
screen "BWTS" 480x228, template "Template_1"
   on GenerateScreen: "TitleUpdater"()
   GraphicView "Graphic view_6" at 70,107 size 332x4; Picture "Graphic_151"
   Button "Button_2" at 88,1 size 50x40; TextOff 'IGGS'
      on Release: ActivateScreen("IGGS Plant", 0)
   Button "Button_4" at 144,1 size 50x40; TextOff 'PGC'
      on Release: ActivateScreen("PGC", 0)
   Button "Button_6" at 199,2 size 50x40; TextOff 'GCU'
      on Release: ActivateScreen("GCU Plant", 0)
   Button "Button_1" at 88,1 size 50x40; TextOff 'IGGS'
      on Release: ActivateScreen("IGGS Plant", 0)
      Visibility <- "IGG Running"
   Button "Button_3" at 144,1 size 50x40; TextOff 'PGC'
      on Release: ActivateScreen("PGC", 0)
      Visibility <- "Process Gas Compressor Running/Stopped"
   Button "Button_5" at 199,2 size 50x40; TextOff 'GCU'
      on Release: ActivateScreen("GCU Plant", 0)
      Visibility <- "100_GCU_AUTO_SEQ_DB_CRNT_STEP"
   Button "HmiScreenItemData_2" at 364,2 size 115x30; TextOn 'I&A Compressor Ok'; TextOff 'Previous Screen'
      on Release: function_efd93a16()
   Button "HmiScreenItemData_19" at 270,2 size 85x40; TextOn 'IGG Plant'; TextOff 'Alarms'
      on Release: ActivateScreen("Alarms", 0)
   Button "Button_20" at 205,191 size 60x34; TextOff 'Dwell'
      Appearance <- "2100_BTCS_CNTRL_DB_BTCS_STATE"
   Button "Button_21" at 2,191 size 60x34; TextOff 'Un- selected'
      Appearance <- "HMI Indication Logic_DB_Tank Selected"
   Button "Button_22" at 69,191 size 60x34; TextOff 'Selected'
      Appearance <- "HMI Indication Logic_DB_Tank Selected"
   Button "Button_23" at 137,191 size 60x34; TextOff 'De-Oxy'
      Appearance <- "2100_BTCS_CNTRL_DB_BTCS_STEP"
   Button "Button_24" at 272,191 size 60x34; TextOff 'Re-Oxy'
      Appearance <- "2100_BTCS_CNTRL_DB_BTCS_STEP"
   Button "Button_25" at 340,191 size 60x34; TextOff 'Post Dwell'
      Appearance <- "2100_BTCS_CNTRL_DB_BTCS_STATE"
   Button "Button_26" at 408,191 size 70x34; TextOff 'Complete'
      Appearance <- "HMI Indication Logic_DB_Sequence Finished"
   TextField "Text field_1" at 185,171 size 116x21; Text 'TANK STATUS'
   Button "Button_28" at 80,49 size 50x55; TextOff 'Tank 6P'
      on Release: function_efd93a16("Tank 6S Status", 0, 0, -1, 2, 1)
   Button "Button_13" at 80,49 size 50x55; TextOff 'Tank 6P'
      on Release: function_efd93a16("Tank 6S Status", 0, 0, -1, 2, 1)
      Appearance <- "2100_BTCS_CNTRL_DB_BTCS_STATE"
      Visibility <- "504_Tank Grouping_DB2020_GROUP of TANK 12"
   Button "Button_29" at 132,49 size 50x55; TextOff 'Tank 5P'
      on Release: function_efd93a16("Tank 5S Status", 0, 0, -1, 2, 1)
   Button "Button_12" at 132,49 size 50x55; TextOff 'Tank 5P'
      on Release: function_efd93a16("Tank 5S Status", 0, 0, -1, 2, 1)
      Appearance <- "2100_BTCS_CNTRL_DB_BTCS_STATE"
      Visibility <- "504_Tank Grouping_DB2020_GROUP of TANK 10"
   Button "Button_30" at 185,49 size 50x55; TextOff 'Tank 4P'
      on Release: function_efd93a16("Tank 4S Status", 0, 0, -1, 2, 1)
   Button "Button_15" at 185,49 size 50x55; TextOff 'Tank 4P'
      on Release: function_efd93a16("Tank 4S Status", 0, 0, -1, 2, 1)
      Appearance <- "2100_BTCS_CNTRL_DB_BTCS_STATE"
      Visibility <- "504_Tank Grouping_DB2020_GROUP of TANK 8"
   Button "Button_31" at 238,49 size 50x55; TextOff 'Tank 3P'
      on Release: function_efd93a16("Tank 3S Status", 0, 0, -1, 2, 1)
   Button "Button_14" at 238,49 size 50x55; TextOff 'Tank 3P'
      on Release: function_efd93a16("Tank 3S Status", 0, 0, -1, 2, 1)
      Appearance <- "2100_BTCS_CNTRL_DB_BTCS_STATE"
      Visibility <- "504_Tank Grouping_DB2020_GROUP of TANK 6"
   Button "Button_32" at 291,49 size 50x55; TextOff 'Tank 2P'
      on Release: function_efd93a16("Tank 2S Status", 0, 0, -1, 2, 1)
   Button "Button_17" at 291,49 size 50x55; TextOff 'Tank 2P'
      on Release: function_efd93a16("Tank 2S Status", 0, 0, -1, 2, 1)
      Appearance <- "2100_BTCS_CNTRL_DB_BTCS_STATE"
      Visibility <- "504_Tank Grouping_DB2020_GROUP of TANK 4"
   Button "Button_33" at 344,49 size 50x55; TextOff 'Tank 1P'
      on Release: function_efd93a16("Tank 1S Status", 0, 0, -1, 2, 1)
   Button "Button_16" at 344,49 size 50x55; TextOff 'Tank 1P'
      on Release: function_efd93a16("Tank 1S Status", 0, 0, -1, 2, 1)
      Appearance <- "2100_BTCS_CNTRL_DB_BTCS_STATE"
      Visibility <- "504_Tank Grouping_DB2020_GROUP of TANK 2"
   Button "Button_34" at 402,82 size 50x55; TextOff 'FP Tank'
      on Release: function_efd93a16("Tank FP Status", 0, 0, -1, 2, 1)
   Button "Button_19" at 402,82 size 50x55; TextOff 'FP Tank'
      on Release: function_efd93a16("Tank FP Status", 0, 0, -1, 2, 1)
      Appearance <- "2100_BTCS_CNTRL_DB_BTCS_STATE"
      Visibility <- "504_Tank Grouping_DB2020_GROUP of TANK 1"
   Button "Button_35" at 22,82 size 50x55; TextOff 'AP Tank'
      on Release: function_efd93a16("Tank AP Status", 0, 0, -1, 2, 1)
   Button "Button_18" at 22,82 size 50x55; TextOff 'AP Tank'
      on Release: function_efd93a16("Tank AP Status", 0, 0, -1, 2, 1)
      Appearance <- "2100_BTCS_CNTRL_DB_BTCS_STATE"
      Visibility <- "504_Tank Grouping_DB2020_GROUP of TANK 14"
   Button "Button_36" at 80,114 size 50x55; TextOff 'Tank 6S'
      on Release: function_efd93a16("Tank 6P Status", 0, 0, -1, 2, 1)
   Button "Button_7" at 80,114 size 50x55; TextOff 'Tank 6S'
      on Release: function_efd93a16("Tank 6P Status", 0, 0, -1, 2, 1)
      Appearance <- "2100_BTCS_CNTRL_DB_BTCS_STATE"
      Visibility <- "504_Tank Grouping_DB2020_GROUP of TANK 13"
   Button "Button_37" at 132,114 size 50x55; TextOff 'Tank 5S'
      on Release: function_efd93a16("Tank 5P Status", 0, 0, -1, 2, 1)
   Button "Button_27" at 132,114 size 50x55; TextOff 'Tank 5S'
      on Release: function_efd93a16("Tank 5P Status", 0, 0, -1, 2, 1)
      Appearance <- "2100_BTCS_CNTRL_DB_BTCS_STATE"
      Visibility <- "504_Tank Grouping_DB2020_GROUP of TANK 11"
   Button "Button_38" at 185,114 size 50x55; TextOff 'Tank 4S'
      on Release: function_efd93a16("Tank 4P Status", 0, 0, -1, 2, 1)
   Button "Button_9" at 185,114 size 50x55; TextOff 'Tank 4S'
      on Release: function_efd93a16("Tank 4P Status", 0, 0, -1, 2, 1)
      Appearance <- "2100_BTCS_CNTRL_DB_BTCS_STATE"
      Visibility <- "504_Tank Grouping_DB2020_GROUP of TANK 9"
   Button "Button_39" at 238,114 size 50x55; TextOff 'Tank 3S'
      on Release: function_efd93a16("Tank 3P Status", 0, 0, -1, 2, 1)
   Button "Button_8" at 238,114 size 50x55; TextOff 'Tank 3S'
      on Release: function_efd93a16("Tank 3P Status", 0, 0, -1, 2, 1)
      Appearance <- "2100_BTCS_CNTRL_DB_BTCS_STATE"
      Visibility <- "504_Tank Grouping_DB2020_GROUP of TANK 7"
   Button "Button_40" at 291,114 size 50x55; TextOff 'Tank 2S'
      on Release: function_efd93a16("Tank 2P Status", 0, 0, -1, 2, 1)
   Button "Button_11" at 291,114 size 50x55; TextOff 'Tank 2S'
      on Release: function_efd93a16("Tank 2P Status", 0, 0, -1, 2, 1)
      Appearance <- "2100_BTCS_CNTRL_DB_BTCS_STATE"
      Visibility <- "504_Tank Grouping_DB2020_GROUP of TANK 5"
   Button "Button_41" at 344,114 size 50x55; TextOff 'Tank 1S'
      on Release: function_efd93a16("Tank 1P Status", 0, 0, -1, 2, 1)
   Button "Button_10" at 344,114 size 50x55; TextOff 'Tank 1S'
      on Release: function_efd93a16("Tank 1P Status", 0, 0, -1, 2, 1)
      Appearance <- "2100_BTCS_CNTRL_DB_BTCS_STATE"
      Visibility <- "504_Tank Grouping_DB2020_GROUP of TANK 3"
   Polyline "Polyline_1" at 80,49 size 48x54
      Visibility <- "504_Tank Grouping_DB2020_RUN TANK 12"
   Polyline "Polyline_2" at 80,114 size 48x54
      Visibility <- "504_Tank Grouping_DB2020_RUN TANK 13"
   Polyline "Polyline_3" at 133,114 size 48x54
      Visibility <- "504_Tank Grouping_DB2020_RUN TANK 11"
   Polyline "Polyline_4" at 132,49 size 48x54
      Visibility <- "504_Tank Grouping_DB2020_RUN TANK 10"
   Polyline "Polyline_5" at 185,49 size 48x54
      Visibility <- "504_Tank Grouping_DB2020_RUN TANK 8"
   Polyline "Polyline_6" at 185,114 size 48x54
      Visibility <- "504_Tank Grouping_DB2020_RUN TANK 9"
   Polyline "Polyline_7" at 239,49 size 48x54
      Visibility <- "504_Tank Grouping_DB2020_RUN TANK 6"
   Polyline "Polyline_8" at 238,114 size 48x54
      Visibility <- "504_Tank Grouping_DB2020_RUN TANK 7"
   Polyline "Polyline_9" at 292,114 size 48x54
      Visibility <- "504_Tank Grouping_DB2020_RUN TANK 5"
   Polyline "Polyline_10" at 291,49 size 48x54
      Visibility <- "504_Tank Grouping_DB2020_RUN TANK 4"
   Polyline "Polyline_11" at 345,49 size 48x54
      Visibility <- "504_Tank Grouping_DB2020_RUN TANK 2"
   Polyline "Polyline_12" at 345,114 size 48x54
      Visibility <- "504_Tank Grouping_DB2020_RUN TANK 3"
   Polyline "Polyline_13" at 403,82 size 48x54
      Visibility <- "504_Tank Grouping_DB2020_RUN TANK 1"
   Polyline "Polyline_14" at 22,82 size 48x54
      Visibility <- "504_Tank Grouping_DB2020_RUN TANK 14"
   Button "HmiScreenItemData_1" at 1,1 size 84x30; TextOn 'I&A Compressor Ok'; TextOff 'Main Index'
      on Release: ActivateScreen("Main Index", 0)

screen "PGC" 480x228, template "Template_1"
   on GenerateScreen: "TitleUpdater"()
   Button "HmiScreenItemData_6" at 353,1 size 126x30; TextOn 'I&A Compressor Ok'; TextOff 'Previous Screen'
      on Release: function_efd93a16()
   TextField "Text field_7" at 4,38 size 278x22; Text 'Process Gas Compressor Control'
   Button "Button_15" at 23,138 size 57x23; TextOn 'Enabled'; TextOff 'Disabled'
   Button "Button_16" at 177,138 size 64x23; TextOn 'Alarm'; TextOff 'Text'
   TextField "Text field_15" at 27,118 size 56x17; Text 'Enabled'
   TextField "Text field_16" at 102,118 size 58x17; Text 'Running'
   TextField "Text field_18" at 179,117 size 69x17; Text 'Shutdown'
   Button "Button_1" at 100,138 size 57x23; TextOn 'Enabled'; TextOff 'Stopped'
   TextField "Text field_32" at 23,139 size 57x23; Text 'Enabled'
      Visibility <- "10_DI_DATA_E_400_SHTDN"
   TextField "Text field_2" at 100,138 size 57x23; Text 'Running'
      Visibility <- "10_DI_DATA_E_400_RUN"
   Button "Button_2" at 177,138 size 64x23; TextOn 'Alarm'; TextOff 'Shutdown'
      Appearance <- "10_DI_DATA_E_400_NOK"
      Visibility <- "10_DI_DATA_E_400_NOK"
   Button "Button_7" at 262,38 size 57x23; TextOn 'Alarm'; TextOff 'Service'
      Appearance <- "140_PGC_HRS_RUN_DB_SRVC"
   GraphicView "Graphic view_1" at 288,29 size 192x199; Picture "Graphic_251"
   Button "HmiScreenItemData_1" at 1,1 size 84x30; TextOn 'I&A Compressor Ok'; TextOff 'Main Index'
      on Release: ActivateScreen("Main Index", 0)

screen "CA Blower" 480x228, template "Template_1"
   on GenerateScreen: "TitleUpdater"()
   Button "HmiScreenItemData_6" at 353,1 size 126x30; TextOn 'I&A Compressor Ok'; TextOff 'Previous Screen'
      on Release: function_efd93a16()
   GraphicIOField "Graphic I/O field_2" at 281,42 size 196x184; PictureList "IA Compressor"
      ProcessValue <- "CA Blower Animation"
   Button "Button_3" at 126,118 size 57x23; TextOn 'Enabled'; TextOff 'Disabled'
   TextField "Text field_4" at 129,98 size 56x17; Text 'Enabled'
   TextField "Text field_5" at 202,98 size 38x17; Text 'Fault'
   Button "Button_5" at 192,118 size 57x23; TextOn 'Enabled'; TextOff 'Healthy'
   TextField "Text field_8" at 126,118 size 57x23; Text 'Enabled'
      Visibility <- "CA Blower Control"
   Button "Button_6" at 192,118 size 57x23; TextOn 'Alarm'; TextOff 'Fault'
      Visibility <- "Data To IGG PLC_Data_VSD Fault Flag"
      Appearance <- "Data To IGG PLC_Data_VSD Fault Flag"
   TextField "Text field_3" at 5,120 size 119x18; Text 'Combustion Air'
   TextField "Text field_7" at 4,38 size 263x22; Text 'Combustion Air Blower Control'
   Button "Button_7" at 276,38 size 57x23; TextOn 'Alarm'; TextOff 'Service'
      Appearance <- "Operation hours E139_IDB_Service Time bit"
   Button "HmiScreenItemData_1" at 1,1 size 84x30; TextOn 'I&A Compressor Ok'; TextOff 'Main Index'
      on Release: ActivateScreen("Main Index", 0)

screen "Cooling System" 480x228, template "Template_1"
   on GenerateScreen: "TitleUpdater"()
   Button "HmiScreenItemData_6" at 353,1 size 126x30; TextOn 'I&A Compressor Ok'; TextOff 'Previous Screen'
      on Release: function_efd93a16()
   TextField "Text field_7" at 140,69 size 201x22; Text 'Cooling System Control'
   Button "Button_15" at 207,128 size 57x23; TextOn 'Enabled'; TextOff 'Disabled'
   Button "Button_16" at 361,128 size 64x23; TextOn 'Alarm'; TextOff 'Text'
   TextField "Text field_14" at 35,130 size 179x18; Text 'Cooling Sea Water Pump'
   TextField "Text field_15" at 211,108 size 56x17; Text 'Enabled'
   TextField "Text field_16" at 286,108 size 58x17; Text 'Running'
   TextField "Text field_18" at 363,107 size 69x17; Text 'Shutdown'
   Rectangle "Rectangle_10" at 33,123 size 166x32
      Appearance <- "P301 Present"
   Button "Button_1" at 284,128 size 57x23; TextOn 'Enabled'; TextOff 'Stopped'
   TextField "Text field_32" at 207,128 size 57x23; Text 'Enabled'
      Visibility <- "CSW Pump Enabled"
   TextField "Text field_2" at 284,128 size 57x23; Text 'Running'
      Visibility <- "Data_To_BC PLC_Data_Cooling Water System Proved"
   Button "Button_2" at 361,128 size 64x23; TextOn 'Alarm'; TextOff 'Shutdown'
      Visibility <- "Cooling Sea Water Pump Shutdown"
      Appearance <- "Cooling Sea Water Pump Shutdown"
   Rectangle "Rectangle_1" at 24,99 size 425x69
      Visibility <- "P301 Present"
   Group "Group" at 15,161 size 490x34
   Button "HmiScreenItemData_1" at 1,1 size 84x30; TextOn 'I&A Compressor Ok'; TextOff 'Main Index'
      on Release: ActivateScreen("Main Index", 0)
   TextField "Text field_1" at 28,161 size 466x34; Text 'Cooling System Pressure in Range'
      Visibility <- "Cooling System Operating"
   TextField "Text field_3" at 15,162 size 490x32; Text 'Cooling System Pressure Out of Range'
      Visibility <- "Cooling System Operating"

screen "Fuel System" 480x228, template "Template_1"
   on GenerateScreen: "TitleUpdater"()
   Button "HmiScreenItemData_6" at 172,1 size 126x30; TextOn 'I&A Compressor Ok'; TextOff 'Previous Screen'
      on Release: function_efd93a16()
   GraphicView "Graphic view_4" at 271,104 size 24x23; Picture "Graphic_102"
   TextField "Text field_3" at 359,196 size 55x18; Text 'E-500B'
   GraphicView "Graphic view_16" at 326,49 size 123x15; Picture "Graphic_99"
   GraphicIOField "Graphic I/O field_1" at 354,30 size 60x65; PictureList "Pump Ani"
      ProcessValue <- "Fuel Pump 1 Animation"
   GraphicView "Graphic view_10" at 325,151 size 124x15; Picture "Graphic_99"
   GraphicIOField "Graphic I/O field_2" at 354,133 size 60x65; PictureList "Pump Ani"
      ProcessValue <- "Fuel Pump 2 Animation"
   GraphicView "Graphic view_17" at 310,64 size 15x94; Picture "Graphic_101"
   GraphicView "Graphic view_14" at 311,140 size 21x25; Picture "Graphic_96"
   GraphicView "Graphic view_18" at 311,50 size 24x23; Picture "Graphic_102"
   GraphicView "Graphic view_19" at 306,99 size 18x23; Picture "Graphic_105"
   GraphicView "Graphic view_20" at 450,64 size 15x94; Picture "Graphic_101"
   GraphicView "Graphic view_9" at 440,50 size 24x23; Picture "Graphic_104"
   GraphicView "Graphic view_21" at 439,141 size 25x24; Picture "Graphic_97"
   GraphicView "Graphic view_7" at 451,100 size 19x24; Picture "Graphic_103"
   GraphicView "Graphic view_22" at 296,103 size 9x15; Picture "Graphic_99"
   GraphicView "Graphic view_24" at 340,49 size 18x15; Picture "Graphic_99"
   TextField "Text field_2" at 359,96 size 56x18; Text 'E-500A'
   GraphicView "Graphic view_1" at 289,103 size 27x15; Picture "Graphic_99"
   Rectangle "Rectangle_13" at 346,24 size 77x92
      Appearance <- "Fuel Pump 1 Tripped"
   Rectangle "Rectangle_14" at 346,127 size 77x92
      Appearance <- "Fuel Pump 2 Tripped"
   TextField "Text field_7" at 334,225 size 83x18; Text 'Duty Pump'
      Visibility <- "101_Fuel_Pumps_DB_Duty Is B"
   TextField "Text field_12" at 346,7 size 83x18; Text 'Duty Pump'
      Visibility <- "101_Fuel_Pumps_DB_Duty Is A"
   Button "HmiScreenItemData_7" at 209,128 size 84x37; TextOn 'Back'; TextOff 'PSelect'; Authorization "Operate"
      on Press: function_b14e0dd5("HMI Fuel Pump Duty Select", 0)
   Button "Button_15" at 7,61 size 57x25; TextOn 'Enabled'; TextOff 'Disabled'
   TextField "Text field_14" at 1,92 size 92x20; Text 'Fuel Pump 1'
   TextField "Text field_15" at 11,40 size 60x18; Text 'Enabled'
   Button "Button_17" at 229,61 size 57x25; TextOn 'Alarm'; TextOff 'Service'
   Button "Button_9" at 229,61 size 57x25; TextOn 'Alarm'; TextOff 'Service'
      Visibility <- "82_To_HMI_E500A Fuel Pump Service Due"
   Button "Button_13" at 7,61 size 57x25; TextOn 'Enabled'; TextOff 'Enabled'
      Visibility <- "Fuel Pump 1 Enabled"
   IOField "I/O field_3" at 131,61 size 65x25; FormatPattern 999999
      ProcessValue <- "64_Functioning Hours_E500A_IDB_Hours Functioning"
   TextField "Text field_5" at 131,38 size 72x18; Text 'Hour Run'
   Button "Button_1" at 70,61 size 57x25; TextOn 'Alarm'; TextOff 'Text'
   TextField "Text field_6" at 78,38 size 45x18; Text 'Alarm'
   Button "Button_3" at 70,61 size 57x25; TextOn 'Alarm'; TextOff 'Tripped'
      Visibility <- "Fuel Pump 1 Tripped"
      Appearance <- "Fuel Pump 1 Tripped"
   Button "Button_18" at 7,178 size 57x25; TextOn 'Enabled'; TextOff 'Disabled'
   TextField "Text field_19" at 1,208 size 92x20; Text 'Fuel Pump 2'
   Button "Button_20" at 229,178 size 57x25; TextOn 'Alarm'; TextOff 'Service'
   Button "Button_10" at 229,178 size 57x25; TextOn 'Alarm'; TextOff 'Service'
      Visibility <- "82_To_HMI_E500B Fuel Pump Service Due"
   Button "Button_14" at 7,177 size 57x25; TextOn 'Enabled'; TextOff 'Enabled'
      Visibility <- "Fuel Pump 2 Enabled"
   IOField "I/O field_6" at 131,177 size 65x25; FormatPattern 999999
      ProcessValue <- "64_Functioning Hours_E500B_IDB_Hours Functioning"
   Button "Button_2" at 70,177 size 57x25; TextOn 'Alarm'; TextOff 'Text'
   Button "Button_4" at 70,177 size 57x25; TextOn 'Alarm'; TextOff 'Tripped'
      Visibility <- "Fuel Pump 2 Tripped"
      Appearance <- "Fuel Pump 2 Tripped"
   Button "HmiScreenItemData_1" at 1,1 size 84x30; TextOn 'I&A Compressor Ok'; TextOff 'Main Index'
      on Release: ActivateScreen("Main Index", 0)

screen "Alarms" 480x228, template "Template_1"
   on GenerateScreen: "TitleUpdater"()
   AlarmView "Alarm view_1" at 0,31 size 480x196
   Button "HmiScreenItemData_6" at 353,1 size 126x30; TextOn 'I&A Compressor Ok'; TextOff 'Previous Screen'
      on Release: function_efd93a16()
   Button "HmiScreenItemData_1" at 1,1 size 84x30; TextOn 'I&A Compressor Ok'; TextOff 'Main Index'
      on Release: ActivateScreen("Main Index", 0)

screen "Events History" 480x228, template "Template_1"
   on GenerateScreen: "TitleUpdater"()
   AlarmView "Alarm view_1" at 0,44 size 480x184
   Button "HmiScreenItemData_1" at 1,1 size 84x30; TextOn 'I&A Compressor Ok'; TextOff 'Main Index'
      on Release: ActivateScreen("Main Index", 0)

screen "Air System" 480x228, template "Template_1"
   on GenerateScreen: "TitleUpdater"()
   Button "HmiScreenItemData_6" at 353,1 size 126x30; TextOn 'I&A Compressor Ok'; TextOff 'Previous Screen'
      on Release: function_efd93a16()
   TextField "Text field_1" at 0,38 size 368x23; Text 'Instrument & Atomising Air Compressor'
   Button "Button_4" at 362,39 size 57x23; TextOn 'Alarm'; TextOff 'Service'
      Visibility <- "IDB_E131_Functioning Hours_Service Time bit"
      Appearance <- "IDB_E131_Functioning Hours_Service Time bit"
   Button "Button_15" at 27,137 size 57x23; TextOn 'Enabled'; TextOff 'Disabled'
   Button "Button_16" at 181,137 size 64x23; TextOn 'Alarm'; TextOff 'Text'
   TextField "Text field_15" at 25,117 size 62x20; Text 'Enabled'
   TextField "Text field_16" at 101,117 size 64x20; Text 'Running'
   TextField "Text field_18" at 174,116 size 78x20; Text 'Shutdown'
   Button "Button_1" at 104,137 size 57x23; TextOn 'Enabled'; TextOff 'Stopped'
   TextField "Text field_32" at 27,137 size 57x23; Text 'Enabled'
      Visibility <- "IA Comp Control"
   TextField "Text field_2" at 104,137 size 57x23; Text 'Running'
      Visibility <- "IA Compressor Healthy"
   Button "Button_2" at 181,137 size 64x23; TextOn 'Alarm'; TextOff 'Shutdown'
      Appearance <- "IA Compressor Shutdown Active"
   GraphicView "Graphic view_91" at 294,85 size 113x127; Picture "Graphic_246"
   GraphicIOField "Graphic I/O field_5" at 286,78 size 129x139; PictureList "New IA Compressor"
      Visibility <- "Data_From BC PLC_Data_IA Compressor Running"
      ProcessValue <- "IA Compressor Animation"
   GraphicView "Graphic view_93" at 419,82 size 48x132; Picture "Graphic_248"
   GraphicView "Graphic view_19" at 404,138 size 19x12; Picture "Graphic_63"
   GraphicView "Graphic view_79" at 404,174 size 19x12; Picture "Graphic_63"
   Bar "Bar_1" at 433,91 size 20x105; Unit  %; MinimumValue 0; MaximumValue 100
      ProcessValue <- "Inlet IA Pressure PIT112 Scaled"
      MaximumValue <- "HMI Data_Inlet IA Pressure (PIT112) High High"
   Button "HmiScreenItemData_1" at 1,1 size 84x30; TextOn 'I&A Compressor Ok'; TextOff 'Main Index'
      on Release: ActivateScreen("Main Index", 0)

Template "Template_1" 480x228
   Softkey "Softkey_F1" at 37,208 size 64x64
      on KeyDown: ActivateScreen("Main Index", 0)
   Softkey "Softkey_F2" at 151,208 size 64x64
      on KeyDown: ActivateScreen("IGGS Plant", 0)
   Softkey "Softkey_F3" at 265,208 size 64x64
      on KeyDown: ActivateScreen("BWTS", 0)
   Softkey "Softkey_F4" at 379,208 size 64x64
      on KeyDown: ActivateScreen("Alarms", 0)
   Circle "Circle_46" at 234,1 size 26x26
      Visibility <- "TRUE"
      Appearance <- "IGG PLC HEART BEAT"
   Circle "Circle_1" at 204,1 size 26x26
      Visibility <- "TRUE"
      Appearance <- "Setpoint Override_DB_Set Pressure"

PopupScreen "Tank 1P Status" 480x272
   TextField "Text field_4" at 9,136 size 86x22; Text 'Pressure:'
   IOField "I/O field_1" at 142,131 size 90x25; FormatPattern s999.9; Unit  mBar
      ProcessValue <- "20_TANKS_IP_DATA_RIO_01_SECOND_TANK_TANKS_PRESS"
   TextField "Text field_5" at 9,170 size 113x22; Text 'Water Level:'
   IOField "I/O field_2" at 142,165 size 90x25; FormatPattern 999.9; Unit  %
      ProcessValue <- "20_TANKS_IP_DATA_RIO_01_SECOND_TANK_BWT_LEVEL"
   TextField "Text field_6" at 9,204 size 137x22; Text 'MBG Flow Rate:'
   IOField "I/O field_3" at 142,199 size 90x25; FormatPattern 999.9; Unit  m³/hr
      ProcessValue <- "20_TANKS_IP_DATA_RIO_01_SECOND_TANK_MBG_FLOW"
   TextField "Text field_7" at 9,238 size 135x22; Text 'USD Flow Rate:'
   IOField "I/O field_4" at 142,233 size 90x25; FormatPattern 999.9; Unit  m³/hr
      ProcessValue <- "20_TANKS_IP_DATA_RIO_01_SECOND_TANK_USD_FLOW"
   Button "Button_1" at 51,5 size 186x35; TextOff 'Port Tank 1 (1P)'
      on Release: function_efd93a16("Tank 1P Status", 0, 0, -1, 0, 1)
   TextField "Text field_1" at 5,90 size 109x25; Text 'TIME LEFT:'
   GraphicView "Graphic view_1" at 9,46 size 223x32; Picture "Tank Manually Disabled"
   GraphicIOField "Graphic I/O field_1" at 9,46 size 223x32; PictureList "Tank Process Stage_II"
      ProcessValue <- "2100_BTCS_CNTRL_DB_BTCS_STATE"
      Visibility <- "504_Tank Grouping_DB2020_GROUP of TANK 2"
   Button "Button_2" at 4,5 size 45x35; TextOff 'Text'; PictureOff "Graphic_286"
      on Click: function_efd93a16("Tank 1P Status", 0, 0, -1, -1, 1)
   IOField "I/O field_29" at 189,90 size 47x25; FormatPattern 99; Unit m
      ProcessValue <- "504_Tank Grouping_DB2020_Time Left Tank_Time Left m Tank 2"
   IOField "I/O field_8" at 146,90 size 42x25; FormatPattern 99; Unit h
      ProcessValue <- "504_Tank Grouping_DB2020_Time Left Tank_Time Left h Tank 2"
   IOField "I/O field_9" at 103,90 size 42x25; FormatPattern 99; Unit d
      ProcessValue <- "504_Tank Grouping_DB2020_Time Left Tank_Time Left d Tank 2"
   TextField "Text field_8" at 235,135 size 140x22; Text 'Water pH Level:'
   IOField "I/O field_5" at 378,130 size 90x25; FormatPattern 99.9
      ProcessValue <- "20_TANKS_IP_DATA_RIO_01_SECOND_TANK_BWT_PH"
   TextField "Text field_9" at 237,170 size 143x22; Text 'Water DO Level:'
   IOField "I/O field_6" at 378,165 size 90x25; FormatPattern 99.99; Unit  mg/l
      ProcessValue <- "20_TANKS_IP_DATA_RIO_01_SECOND_TANK_BWT_DO"
   TextField "Text field_10" at 236,204 size 174x22; Text 'Water Temperature:'
   IOField "I/O field_7" at 393,199 size 75x25; FormatPattern 999.9; Unit  °C
      ProcessValue <- "20_TANKS_IP_DATA_RIO_01_SECOND_TANK_BWT_TEMP"
   Group "Group" at 242,229 size 225x40; Authorization "Operate"
   Button "Button_5" at 242,229 size 225x40; TextOff 'Tank Shutdown Alarm'
      Visibility <- "2062_Warning_Data_Alarm Tank P1"
      ProcessValue <- "2062_Warning_Data_Water Level Override 1P"
   Button "Button_6" at 242,229 size 225x40; TextOff 'No/Low Water Level'; Authorization "Operate"
      ProcessValue <- "2062_Warning_Data_Water Level Override 1P"
      Visibility <- "LT422 1P  TANK LEVEL ALARM_ALARM L"